            Reaction_time_after_command : Bool := TRUE;   // Start reaction time after command or after shotend
            Spare_0_2 : Bool := FALSE;
            Spare_0_3 : Bool := FALSE;
            Spare_0_4 : Bool := FALSE;
            Spare_0_5 : Bool := FALSE;
            Spare_0_6 : Bool := FALSE;
            Spare_0_7 : Bool := FALSE;
            Spare_1_0 : Bool := FALSE;
            Spare_1_1 : Bool := FALSE;
            Spare_1_2 : Bool := FALSE;
            Spare_1_3 : Bool := FALSE;
            Spare_1_4 : Bool := FALSE;
            Spare_1_5 : Bool := FALSE;
            Spare_1_6 : Bool := FALSE;
            Spare_1_7 : Bool := FALSE;
            Spare_2_0 : Bool := FALSE;
            Spare_2_1 : Bool := FALSE;
            Vacuum_button_valve_1 : Bool := FALSE;
            Vacuum_button_valve_2 : Bool := FALSE;
            Vacuum_button_valve_3 : Bool := TRUE;
            Vacuum_button_valve_4 : Bool := FALSE;
            Vacuum_button_valve_5 : Bool := FALSE;
            Vacuum_button_valve_6 : Bool := FALSE;
            Spare_3 : Byte := 16#00;
         END_STRUCT;
         Times_WinCap : Struct
            SOD_core_WP : Array[0..32] of Time;   // switch on delay core WP
            SOD_core_BP : Array[0..32] of Time;   // switch on delay core BP
            Duration_core : Array[0..32] of Time;   // duration core without endposition
         END_STRUCT;
         Settings_Special : Struct
            Config_write : Bool := FALSE;
            Config_write_done : Bool := FALSE;
            Spare : Int := 1;
            Core_Input : Array[0..32] of "UDT_CoreSettingsSpecial";
            Core_Type : Array[0..32] of Struct
               NC_WP_1 : Bool;   // Schließerkontakt = 0
               NC_WP_2 : Bool;   // Schließerkontakt = 0
               NC_WP_3 : Bool;   // Schließerkontakt = 0
               NC_WP_4 : Bool;   // Schließerkontakt = 0
               NC_WP_5 : Bool;   // Schließerkontakt = 0
               NC_WP_6 : Bool;   // Schließerkontakt = 0
               Forced_forward_WP : Bool;   // Dauernd angesteuert
               Signal_from_upper_tool_WP : Bool;
               NC_BP_1 : Bool;   // Schließerkontakt = 0
               NC_BP_2 : Bool;   // Schließerkontakt = 0
               NC_BP_3 : Bool;   // Schließerkontakt = 0
               NC_BP_4 : Bool;   // Schließerkontakt = 0
               NC_BP_5 : Bool;   // Schließerkontakt = 0
               NC_BP_6 : Bool;   // Schließerkontakt = 0
               Forced_forward_BP : Bool;   // Dauernd angesteuert
               Signal_from_upper_tool_BP : Bool;
            END_STRUCT;
            Config_I_O : Struct
               Lower_tool_card : Array[1..16] of Bool;   // Karte vorhanden
               Upper_tool_card : Array[1..16] of Bool;   // Karte vorhanden
            END_STRUCT;
         END_STRUCT;
      END_STRUCT;
      Set_flow_seals : Struct
         Warning_Tolerance : Struct   // Warning/Tolerance for each seal
            Warning : Array[0..32] of Int;
            Tolerance : Array[0..32] of Int;
         END_STRUCT;
         Set_flow : Array[0..32] of Int;
         Warning_all : Int;   // Warning for all seals
         Tolerance_all : Int;   // Tolerance for all seals
         Set_flow_all : Int;
         Offset_Flow_1 : Real;
         Offset_Flow_2 : Real;
         Offset_Flow_3 : Real;
         SOD_Seal_test : Time := T#2S;   // Waittime to check seal flow
         Spare_140 : Int;
         Spare_142 : Int;
         Spare_144 : Int;
         Spare_146 : Int;
      END_STRUCT;
   END_STRUCT;
   // Set_times_movement.Time_MC_WP[0] := T#10S;
   // Set_times_movement.Time_MC_WP[1] := T#10S;
   // Set_times_movement.Time_MC_WP[2] := T#10S;
   // Set_times_movement.Time_MC_WP[3] := T#10S;
   // Set_times_movement.Time_MC_WP[4] := T#10S;
   // Set_times_movement.Time_MC_WP[5] := T#10S;
   // Set_times_movement.Time_MC_WP[6] := T#10S;
   // Set_times_movement.Time_MC_WP[7] := T#10S;
   // Set_times_movement.Time_MC_WP[8] := T#10S;
   // Set_times_movement.Time_MC_WP[9] := T#10S;
   // Set_times_movement.Time_MC_WP[10] := T#10S;
   // Set_times_movement.Time_MC_WP[11] := T#10S;
   // Set_times_movement.Time_MC_WP[12] := T#10S;
   // Set_times_movement.Time_MC_WP[13] := T#10S;
   // Set_times_movement.Time_MC_WP[14] := T#10S;
   // Set_times_movement.Time_MC_WP[15] := T#10S;
   // Set_times_movement.Time_MC_WP[16] := T#10S;
   // Set_times_movement.Time_MC_WP[17] := T#10S;
   // Set_times_movement.Time_MC_WP[18] := T#10S;
   // Set_times_movement.Time_MC_WP[19] := T#10S;
   // Set_times_movement.Time_MC_WP[20] := T#10S;
   // Set_times_movement.Time_MC_WP[21] := T#10S;
   // Set_times_movement.Time_MC_WP[22] := T#10S;
   // Set_times_movement.Time_MC_WP[23] := T#10S;
   // Set_times_movement.Time_MC_WP[24] := T#10S;
   // Set_times_movement.Time_MC_WP[25] := T#10S;
   // Set_times_movement.Time_MC_WP[26] := T#10S;
   // Set_times_movement.Time_MC_WP[27] := T#10S;
   // Set_times_movement.Time_MC_WP[28] := T#10S;
   // Set_times_movement.Time_MC_WP[29] := T#10S;
   // Set_times_movement.Time_MC_WP[30] := T#10S;
   // Set_times_movement.Time_MC_WP[31] := T#10S;
   // Set_times_movement.Time_MC_WP[32] := T#10S;
   // Set_times_movement.Time_MC_BP[0] := T#10S;
   // Set_times_movement.Time_MC_BP[1] := T#10S;
   // Set_times_movement.Time_MC_BP[2] := T#10S;
   // Set_times_movement.Time_MC_BP[3] := T#10S;
   // Set_times_movement.Time_MC_BP[4] := T#10S;
   // Set_times_movement.Time_MC_BP[5] := T#10S;
   // Set_times_movement.Time_MC_BP[6] := T#10S;
   // Set_times_movement.Time_MC_BP[7] := T#10S;
   // Set_times_movement.Time_MC_BP[8] := T#10S;
   // Set_times_movement.Time_MC_BP[9] := T#10S;
   // Set_times_movement.Time_MC_BP[10] := T#10S;
   // Set_times_movement.Time_MC_BP[11] := T#10S;
   // Set_times_movement.Time_MC_BP[12] := T#10S;
   // Set_times_movement.Time_MC_BP[13] := T#10S;
   // Set_times_movement.Time_MC_BP[14] := T#10S;
   // Set_times_movement.Time_MC_BP[15] := T#10S;
   // Set_times_movement.Time_MC_BP[16] := T#10S;
   // Set_times_movement.Time_MC_BP[17] := T#10S;
   // Set_times_movement.Time_MC_BP[18] := T#10S;
   // Set_times_movement.Time_MC_BP[19] := T#10S;
   // Set_times_movement.Time_MC_BP[20] := T#10S;
   // Set_times_movement.Time_MC_BP[21] := T#10S;
   // Set_times_movement.Time_MC_BP[22] := T#10S;
   // Set_times_movement.Time_MC_BP[23] := T#10S;
   // Set_times_movement.Time_MC_BP[24] := T#10S;
   // Set_times_movement.Time_MC_BP[25] := T#10S;
   // Set_times_movement.Time_MC_BP[26] := T#10S;
   // Set_times_movement.Time_MC_BP[27] := T#10S;
   // Set_times_movement.Time_MC_BP[28] := T#10S;
   // Set_times_movement.Time_MC_BP[29] := T#10S;
   // Set_times_movement.Time_MC_BP[30] := T#10S;
   // Set_times_movement.Time_MC_BP[31] := T#10S;
   // Set_times_movement.Time_MC_BP[32] := T#10S;
   // Set_times_movement.Time_MLD_WP[0] := T#10S;
   // Set_times_movement.Time_MLD_WP[1] := T#10S;
   // Set_times_movement.Time_MLD_WP[2] := T#10S;
   // Set_times_movement.Time_MLD_WP[3] := T#10S;
   // Set_times_movement.Time_MLD_WP[4] := T#10S;
   // Set_times_movement.Time_MLD_WP[5] := T#10S;
   // Set_times_movement.Time_MLD_WP[6] := T#10S;
   // Set_times_movement.Time_MLD_WP[7] := T#10S;
   // Set_times_movement.Time_MLD_WP[8] := T#10S;
   // Set_times_movement.Time_MLD_WP[9] := T#10S;
   // Set_times_movement.Time_MLD_WP[10] := T#10S;
   // Set_times_movement.Time_MLD_WP[11] := T#10S;
   // Set_times_movement.Time_MLD_WP[12] := T#10S;
   // Set_times_movement.Time_MLD_WP[13] := T#10S;
   // Set_times_movement.Time_MLD_WP[14] := T#10S;
   // Set_times_movement.Time_MLD_WP[15] := T#10S;
   // Set_times_movement.Time_MLD_WP[16] := T#10S;
   // Set_times_movement.Time_MLD_WP[17] := T#10S;
   // Set_times_movement.Time_MLD_WP[18] := T#10S;
   // Set_times_movement.Time_MLD_WP[19] := T#10S;
   // Set_times_movement.Time_MLD_WP[20] := T#10S;
   // Set_times_movement.Time_MLD_WP[21] := T#10S;
   // Set_times_movement.Time_MLD_WP[22] := T#10S;
   // Set_times_movement.Time_MLD_WP[23] := T#10S;
   // Set_times_movement.Time_MLD_WP[24] := T#10S;
   // Set_times_movement.Time_MLD_WP[25] := T#10S;
   // Set_times_movement.Time_MLD_WP[26] := T#10S;
   // Set_times_movement.Time_MLD_WP[27] := T#10S;
   // Set_times_movement.Time_MLD_WP[28] := T#10S;
   // Set_times_movement.Time_MLD_WP[29] := T#10S;
   // Set_times_movement.Time_MLD_WP[30] := T#10S;
   // Set_times_movement.Time_MLD_WP[31] := T#10S;
   // Set_times_movement.Time_MLD_WP[32] := T#10S;
   // Set_times_movement.Time_MLD_BP[0] := T#10S;
   // Set_times_movement.Time_MLD_BP[1] := T#10S;
   // Set_times_movement.Time_MLD_BP[2] := T#10S;
   // Set_times_movement.Time_MLD_BP[3] := T#10S;
   // Set_times_movement.Time_MLD_BP[4] := T#10S;
   // Set_times_movement.Time_MLD_BP[5] := T#10S;
   // Set_times_movement.Time_MLD_BP[6] := T#10S;
   // Set_times_movement.Time_MLD_BP[7] := T#10S;
   // Set_times_movement.Time_MLD_BP[8] := T#10S;
   // Set_times_movement.Time_MLD_BP[9] := T#10S;
   // Set_times_movement.Time_MLD_BP[10] := T#10S;
   // Set_times_movement.Time_MLD_BP[11] := T#10S;
   // Set_times_movement.Time_MLD_BP[12] := T#10S;
   // Set_times_movement.Time_MLD_BP[13] := T#10S;
   // Set_times_movement.Time_MLD_BP[14] := T#10S;
   // Set_times_movement.Time_MLD_BP[15] := T#10S;
   // Set_times_movement.Time_MLD_BP[16] := T#10S;
   // Set_times_movement.Time_MLD_BP[17] := T#10S;
   // Set_times_movement.Time_MLD_BP[18] := T#10S;
   // Set_times_movement.Time_MLD_BP[19] := T#10S;
   // Set_times_movement.Time_MLD_BP[20] := T#10S;
   // Set_times_movement.Time_MLD_BP[21] := T#10S;
   // Set_times_movement.Time_MLD_BP[22] := T#10S;
   // Set_times_movement.Time_MLD_BP[23] := T#10S;
   // Set_times_movement.Time_MLD_BP[24] := T#10S;
   // Set_times_movement.Time_MLD_BP[25] := T#10S;
   // Set_times_movement.Time_MLD_BP[26] := T#10S;
   // Set_times_movement.Time_MLD_BP[27] := T#10S;
   // Set_times_movement.Time_MLD_BP[28] := T#10S;
   // Set_times_movement.Time_MLD_BP[29] := T#10S;
   // Set_times_movement.Time_MLD_BP[30] := T#10S;
   // Set_times_movement.Time_MLD_BP[31] := T#10S;
   // Set_times_movement.Time_MLD_BP[32] := T#10S;
   // Set_times_seals.SOD_seal[0] := T#2S;
   // Set_times_seals.SOD_seal[1] := T#2S;
   // Set_times_seals.SOD_seal[2] := T#2S;
   // Set_times_seals.SOD_seal[3] := T#2S;
   // Set_times_seals.SOD_seal[4] := T#2S;
   // Set_times_seals.SOD_seal[5] := T#2S;
   // Set_times_seals.SOD_seal[6] := T#2S;
   // Set_times_seals.SOD_seal[7] := T#2S;
   // Set_times_seals.SOD_seal[8] := T#2S;
   // Set_times_seals.SOD_seal[9] := T#2S;
   // Set_times_seals.SOD_seal[10] := T#2S;
   // Set_times_seals.SOD_seal[11] := T#2S;
   // Set_times_seals.SOD_seal[12] := T#2S;
   // Set_times_seals.SOD_seal[13] := T#2S;
   // Set_times_seals.SOD_seal[14] := T#2S;
   // Set_times_seals.SOD_seal[15] := T#2S;
   // Set_times_seals.SOD_seal[16] := T#2S;
   // Set_times_seals.SOD_seal[17] := T#2S;
   // Set_times_seals.SOD_seal[18] := T#2S;
   // Set_times_seals.SOD_seal[19] := T#2S;
   // Set_times_seals.SOD_seal[20] := T#2S;
   // Set_times_seals.SOD_seal[21] := T#2S;
   // Set_times_seals.SOD_seal[22] := T#2S;
   // Set_times_seals.SOD_seal[23] := T#2S;
   // Set_times_seals.SOD_seal[24] := T#2S;
   // Set_times_seals.SOD_seal[25] := T#2S;
   // Set_times_seals.SOD_seal[26] := T#2S;
   // Set_times_seals.SOD_seal[27] := T#2S;
   // Set_times_seals.SOD_seal[28] := T#2S;
   // Set_times_seals.SOD_seal[29] := T#2S;
   // Set_times_seals.SOD_seal[30] := T#2S;
   // Set_times_seals.SOD_seal[31] := T#2S;
   // Set_times_seals.SOD_seal[32] := T#2S;
   // Set_times_seals.Duration_seal[0] := T#1M_1S;
   // Set_times_seals.Duration_seal[1] := T#1M_1S;
   // Set_times_seals.Duration_seal[2] := T#1M;
   // Set_times_seals.Duration_seal[3] := T#1M;
   // Set_times_seals.Duration_seal[4] := T#1M;
   // Set_times_seals.Duration_seal[5] := T#1M;
   // Set_times_seals.Duration_seal[6] := T#1M;
   // Set_times_seals.Duration_seal[7] := T#1M;
   // Set_times_seals.Duration_seal[8] := T#1M;
   // Set_times_seals.Duration_seal[9] := T#1M;
   // Set_times_seals.Duration_seal[10] := T#1M;
   // Set_times_seals.Duration_seal[11] := T#1M;
   // Set_times_seals.Duration_seal[12] := T#1M;
   // Set_times_seals.Duration_seal[13] := T#1M;
   // Set_times_seals.Duration_seal[14] := T#1M;
   // Set_times_seals.Duration_seal[15] := T#1M;
   // Set_times_seals.Duration_seal[16] := T#1M;
   // Set_times_seals.Duration_seal[17] := T#1M;
   // Set_times_seals.Duration_seal[18] := T#1M;
   // Set_times_seals.Duration_seal[19] := T#1M;
   // Set_times_seals.Duration_seal[20] := T#1M;
   // Set_times_seals.Duration_seal[21] := T#1M;
   // Set_times_seals.Duration_seal[22] := T#1M;
   // Set_times_seals.Duration_seal[23] := T#1M;
   // Set_times_seals.Duration_seal[24] := T#1M;
   // Set_times_seals.Duration_seal[25] := T#1M;
   // Set_times_seals.Duration_seal[26] := T#1M;
   // Set_times_seals.Duration_seal[27] := T#1M;
   // Set_times_seals.Duration_seal[28] := T#1M;
   // Set_times_seals.Duration_seal[29] := T#1M;
   // Set_times_seals.Duration_seal[30] := T#1M;
   // Set_times_seals.Duration_seal[31] := T#1M;
   // Set_times_seals.Duration_seal[32] := T#10S;
   // Set_temperature.Setvalue[0] := 0;
   // Set_temperature.Setvalue[1] := 500;
   // // 1726 more start values not shown
END_TYPE

TYPE "UDT_Mould_functions_1"
VERSION : 0.1
   STRUCT
      MouldMovement01WP : Bool;   // 65: Pusher Windshield WP
      MouldMovement02WP : Bool;   // 66: Pusher Knee Border WP
      MouldMovement03WP : Bool;   // 67: Pusher Frontal Area WP
      MouldMovement04WP : Bool;   // 68: Ejector WP
      MouldMovement05WP : Bool;   // 69: Pusher Stössel WP
      MouldMovement06WP : Bool;   // 70: Flip-Flap WP
      MouldMovement07WP : Bool;   // 71: Safty Locking Knee WP
      MouldMovement08WP : Bool;   // 72: Safty Locking WS WP
      MouldMovement09WP : Bool;   // 73: Vacuum lower mould WP
      MouldMovement10WP : Bool;   // 74: Pusher Airbag WP
      MouldMovement11WP : Bool;   // 75: Pusher DS&PS upper mould WP
      MouldMovement12WP : Bool;   // 76: Vacuum upper mould WP
      MouldMovement13WP : Bool;   // 77: Sensor substrate WP
      MouldMovement14WP : Bool;   // 78: Sensor substrate flamed WP
      MouldMovement15WP : Bool;   // 79: Kernzug 15 AS
      MouldMovement16WP : Bool;   // 80: Kernzug 16 AS
      MouldMovement17WP : Bool;   // 81: Kernzug 17 AS
      MouldMovement18WP : Bool;   // 82: Kernzug 18 AS
      MouldMovement19WP : Bool;   // 83: Kernzug 19 AS
      MouldMovement20WP : Bool;   // 84: Kernzug 20 AS
      MouldMovement21WP : Bool;   // 85: Kernzug 21 AS
      MouldMovement22WP : Bool;   // 86: Kernzug 22 AS
      MouldMovement23WP : Bool;   // 87: Kernzug 23 AS
      MouldMovement24WP : Bool;   // 88: Kernzug 24 AS
      MouldMovement25WP : Bool;   // 89: Kernzug 25 AS
      MouldMovement26WP : Bool;   // 90: Kernzug 26 AS
      MouldMovement27WP : Bool;   // 91: Kernzug 27 AS
      MouldMovement28WP : Bool;   // 92: Kernzug 28 AS
      MouldMovement29WP : Bool;   // 93: Kernzug 29 AS
      MouldMovement30WP : Bool;   // 94: Kernzug 30 AS
      MouldMovement31WP : Bool;   // 95: Kernzug 31 AS
      MouldMovement32WP : Bool;   // 96: Kernzug 32 AS
      MouldMovement01BP : Bool;   // 97: Pusher Windshield BP
      MouldMovement02BP : Bool;   // 98: Pusher Knee Border DS BP
      MouldMovement03BP : Bool;   // 99: Pusher Frontal Area BP
      MouldMovement04BP : Bool;   // 100: Ejector BP
      MouldMovement05BP : Bool;   // 101: Pusher Stössel BP
      MouldMovement06BP : Bool;   // 102: Flip-Flap BP
      MouldMovement07BP : Bool;   // 103: Safty Locking Knee BP
      MouldMovement08BP : Bool;   // 104: Safty Locking WS BP
      MouldMovement09BP : Bool;   // 105: Vacuum lower mould BP
      MouldMovement10BP : Bool;   // 106: Pusher Airbag BP
      MouldMovement11BP : Bool;   // 107: Pusher DS&PS upper mould BP
      MouldMovement12BP : Bool;   // 108: Vacuum upper mould BP
      MouldMovement13BP : Bool;   // 109: Sensor substrate BP
      MouldMovement14BP : Bool;   // 110: Sensor substrate flamed BP
      MouldMovement15BP : Bool;   // 111: Kernzug 15 GS
      MouldMovement16BP : Bool;   // 112: Kernzug 16 GS
      MouldMovement17BP : Bool;   // 113: Kernzug 17 GS
      MouldMovement18BP : Bool;   // 114: Kernzug 18 GS
      MouldMovement19BP : Bool;   // 115: Kernzug 19 GS
      MouldMovement20BP : Bool;   // 116: Kernzug 20 GS
      MouldMovement21BP : Bool;   // 117: Kernzug 21 GS
      MouldMovement22BP : Bool;   // 118: Kernzug 22 GS
      MouldMovement23BP : Bool;   // 119: Kernzug 23 GS
      MouldMovement24BP : Bool;   // 120: Kernzug 24 GS
      MouldMovement25BP : Bool;   // 121: Kernzug 25 GS
      MouldMovement26BP : Bool;   // 122: Kernzug 26 GS
      MouldMovement27BP : Bool;   // 123: Kernzug 27 GS
      MouldMovement28BP : Bool;   // 124: Kernzug 28 GS
      MouldMovement29BP : Bool;   // 125: Kernzug 29 GS
      MouldMovement30BP : Bool;   // 126: Kernzug 30 GS
      MouldMovement31BP : Bool;   // 127: Kernzug 31 GS
      MouldMovement32BP : Bool;   // 128: Kernzug 32 GS
   END_STRUCT;
END_TYPE

TYPE "UDT_Tool_Inputs_type_1"
VERSION : 0.1
   STRUCT
      "Lower Mould" : Struct
         "2A1" : Struct
            I_Pusher_Windshield_DS_WP : Bool := FALSE;   // 0.0
            I_Pusher_Windshield_DS_BP : Bool := FALSE;   // 0.1
            Reserve_5 : Bool := FALSE;   // 0.2
            Reserve_4 : Bool := FALSE;   // 0.3
            I_Pusher_Knee_Border_DS_WP : Bool := FALSE;   // 0.4
            I_Pusher_Knee_Border_DS_BP : Bool := FALSE;   // 0.5
            Reserve_3 : Bool := FALSE;   // 0.6
            Reserve_2 : Bool := FALSE;   // 0.7
            I_Pusher_Frontal_Area_DS_WP : Bool := FALSE;   // 1.0
            I_Pusher_Frontal_Area_DS_BP : Bool := FALSE;   // 1.1
            I_Pusher_Frontal_Area_PS_WP : Bool := FALSE;   // 1.2
            I_Pusher_Frontal_Area_PS_BP : Bool := FALSE;   // 1.3
            I_Ejector_WP : Bool := FALSE;   // 1.4
            I_Ejector_BP : Bool := FALSE;   // 1.5
            "I_Flip-Flap_WP" : Bool := FALSE;   // 1.6
            Reserve_1 : Bool := FALSE;   // 1.7
         END_STRUCT;
         "2A2" : Struct
            I_Safty_Locking_Knee_DS_WP : Bool := FALSE;   // 0.0
            I_Safty_Locking_Knee_DS_BP : Bool := FALSE;   // 0.1
            I_Safty_Locking_Knee_PS_WP : Bool := FALSE;   // 0.2
            I_Safty_Locking_Knee_PS_BP : Bool := FALSE;   // 0.3
            I_Safty_Locking_WS_DS_WP : Bool := FALSE;   // 0.4
            I_Safty_Locking_WS_DS_BP : Bool := FALSE;   // 0.5
            I_Safty_Locking_WS_PS_WP : Bool := FALSE;   // 0.6
            I_Safty_Locking_WS_PS_BP : Bool := FALSE;   // 0.7
            "I_Vacuum monitor" : Bool := FALSE;   // 1.0
            Element_2 : Bool := FALSE;   // 1.1
            Element_1 : Bool := FALSE;   // 1.2
            Element_4 : Bool := FALSE;   // 1.3
            Reserve_2 : Bool := FALSE;   // 1.4
            Reserve_3 : Bool := FALSE;   // 1.5
            Reserve_4 : Bool := FALSE;   // 1.6
            Reserve_5 : Bool := FALSE;   // 1.7
         END_STRUCT;
         "2A3" : Struct
            I_Palm_Switch_Vacuum_on : Bool := FALSE;   // 0.0
            I_Illuminated_Key_Vacuum1_off : Bool := FALSE;   // 0.1
            I_Illuminated_Key_Vacuum2_off : Bool := FALSE;   // 0.2
            I_Illuminated_Key_Vacuum3_off : Bool := FALSE;   // 0.3
            Element_3 : Bool := FALSE;   // 0.4
            Element_1 : Bool := FALSE;   // 0.5
            I_PB_Seal_Test_2bar : Bool := FALSE;   // 0.6
            I_2_Hand_active : Bool := FALSE;   // 0.7
            "I_Code_Bit1_(1)" : Bool := FALSE;   // 1.0
            "I_Code_Bit2_(2)" : Bool := FALSE;   // 1.1
            "I_Code_Bit3_(4)" : Bool := FALSE;   // 1.2
            "I_Code_Bit4_(8)" : Bool := FALSE;   // 1.3
            "I_Code_Bit5_(16)" : Bool := FALSE;   // 1.4
            "I_Code_Bit6_(32)" : Bool := FALSE;   // 1.5
            "I_Code_Bit7_(64)" : Bool := FALSE;   // 1.6
            "I_Code_Bit8_(128)" : Bool := FALSE;   // 1.7
         END_STRUCT;
      END_STRUCT;
      "Upper Mould" : Struct
         "46A1" : Struct
            I_Pusher_Airbag_WP : Bool := FALSE;   // 0.0
            I_Pusher_Airbag_BP : Bool := FALSE;   // 0.1
            I_Pusher_DS_WP : Bool := FALSE;   // 0.2
            I_Pusher_DS_BP : Bool := FALSE;   // 0.3
            I_Pusher_PS_WP : Bool := FALSE;   // 0.4
            I_Pusher_PS_BP : Bool := FALSE;   // 0.5
            Element_1 : Bool := FALSE;   // 0.6
            Element_2 : Bool := FALSE;   // 0.7
            I_Vacuum_Motitor : Bool := FALSE;   // 1.0
            I_Sensor_insert : Bool := FALSE;   // 1.1
            I_Sensor_flamed : Bool := FALSE;   // 1.2
            "I_Illuminated Key_Vacuum_off" : Bool := FALSE;   // 1.3
            Element_3 : Bool := FALSE;   // 1.4
            Element_4 : Bool := FALSE;   // 1.5
            Reserve_54 : Bool := FALSE;   // 1.6
            Reserve_55 : Bool := FALSE;   // 1.7
         END_STRUCT;
      END_STRUCT;
   END_STRUCT;
END_TYPE

TYPE "UDT1500_ShotResultToMC"
VERSION : 0.1
   STRUCT
      Data_from_MC : Struct
         Struct01 : Struct
            Data_read : Bool;   // Mouldcarrier has read the shot data
            SPARE_00 : Bool;
            SPARE_01 : Bool;
            SPARE_02 : Bool;
            SPARE_03 : Bool;
            SPARE_04 : Bool;
            SPARE_05 : Bool;
            SPARE_06 : Bool;
            SPARE_07 : Bool;
            SPARE_08 : Bool;
            SPARE_09 : Bool;
            SPARE_10 : Bool;
            SPARE_11 : Bool;
            SPARE_12 : Bool;
            SPARE_13 : Bool;
            SPARE_14 : Bool;
         END_STRUCT;
      END_STRUCT;
      Date_to_MC : Struct
         Struct01 : Struct   // 128 Byte Bereich
            New_Data : Bool;   // Shot Data is now available
            SPARE_00 : Bool;
            SPARE_01 : Bool;
            SPARE_02 : Bool;
            SPARE_03 : Bool;
            SPARE_04 : Bool;
            SPARE_05 : Bool;
            SPARE_06 : Bool;
            FLT_Shottime : Bool;   // Shottime is outside of the tolerance
            FLT_Flowrate_C1 : Bool;   // Flowrate of C1 is outside of the tolerance
            FLT_Flowrate_C2 : Bool;   // Flowrate of C2 is outside of the tolerance
            FLT_PressureMH_C1 : Bool;   // Pressure of C1 at the MH is outside of the tolerance
            FLT_PressureMH_C2 : Bool;   // Pressure of C2 at the MH is outside of the tolerance
            FLT_TempMH_C1 : Bool;   // Temperature of C1 at the MH is outside of the tolerance
            FLT_TempMH_C2 : Bool;   // Temperature of C2 at the MH is outside of the tolerance
            FLT_TempTank_C1 : Bool;   // Temperature of C1 at the tank is outside of the tolerance
            FLT_TempTank_C2 : Bool;   // Temperature of C2 at the tank is outside of the tolerance
            SPARE_07 : Bool;
            SPARE_08 : Bool;
            SPARE_09 : Bool;
            SPARE_10 : Bool;
            SPARE_11 : Bool;
            SPARE_12 : Bool;
            SPARE_13 : Bool;
            SPARE_14 : Bool;
            SPARE_15 : Bool;
            SPARE_16 : Bool;
            SPARE_17 : Bool;
            SPARE_18 : Bool;
            SPARE_19 : Bool;
            SPARE_20 : Bool;
            SPARE_21 : Bool;
            MH_No : Int;   // Number of the MH at the last shot (1 - 16)
            Foam_No : Int;   // Number of foaming program at the last shot (1 - 1000)
            MC_No : Int;
            SPARE_22 : Int;
            Rob_MoveTime : DInt;   // Moving - time of the roboter (1/1 [ms])
            ShotTime_Tol_plus : DInt;   // Tolerance of the shottime (plus) at the last shot (1/1 [ms])
            ShotTime_Setvalue : DInt;   // Setvalue of the shottime at the last shot (1/1 [ms])
            ShotTime_Actvalue : DInt;   // Actual value of the shottime at the last shot (1/1 [ms])
            ShotTime_Tol_minus : DInt;   // Tolerance of the shottime (minus) at the last shot (1/1 [ms])
            ShotWeight_Setvalue : DInt;
            ShotWeight_Actvalue : DInt;
            Flowrate_C1_Tol_plus : DInt;   // Tolerance of the flowrate (plus) at the last shot (1/10 [g/s])
            Flowrate_C1_Setvalue : DInt;   // Setvalue of the flowrate at the last shot (1/10 [g/s])
            Flowrate_C1_Actvalue : DInt;   // Actual value of the flowrate at the last shot (1/10 [g/s])
            Flowrate_C1_Tol_minus : DInt;   // Tolerance of the flowrate (minus) at the last shot (1/10 [g/s])
            Flowrate_C2_Tol_plus : DInt;   // Tolerance of the flowrate (plus) at the last shot (1/10 [g/s])
            Flowrate_C2_Setvalue : DInt;   // Setvalue of the flowrate at the last shot (1/10 [g/s])
            Flowrate_C2_Actvalue : DInt;   // Actual value of the flowrate at the last shot (1/10 [g/s])
            Flowrate_C2_Tol_minus : DInt;   // Tolerance of the flowrate (minus) at the last shot (1/10 [g/s])
            PressureMH_C1_Tol_plus : DInt;   // Tolerance of the pressure of C1 at the MH (plus) at the last shot (1/10 [bar])
            PressureMH_C1_Setvalue : DInt;   // Setvalue of the pressure of C1 at the MH at the last shot (1/10 [bar])
            PressureMH_C1_Actvalue : DInt;   // Actual value of the pressure of C1 at the MH at the last shot (1/10 [bar])
            PressureMH_C1_Tol_minus : DInt;   // Tolerance of the pressure of C1 at the MH(minus) at the last shot (1/10 [bar])
            PressureMH_C2_Tol_plus : DInt;   // Tolerance of the pressure of C2 at the MH (plus) at the last shot (1/10 [bar])
            PressureMH_C2_Setvalue : DInt;   // Setvalue of the pressure of C2 at the MH at the last shot (1/10 [bar])
            PressureMH_C2_Actvalue : DInt;   // Actual value of the pressure of C2 at the MH at the last shot (1/10 [bar])
            PressureMH_C2_Tol_minus : DInt;   // Tolerance of the pressure of C2 at the MH(minus) at the last shot (1/10 [bar])
            TempMH_C1_Tol_plus : DInt;   // Tolerance of the temp. of C1 at the MH (plus) at the last shot (1/10 [°C])
            TempMH_C1_Setvalue : DInt;   // Setvalue of the temp. of C1 at the MH at the last shot (1/10 [°C])
            TempMH_C1_Actvalue : DInt;   // Actual value of the temp. of C1 at the MH at the last shot (1/10 [°C])
            TempMH_C1_Tol_minus : DInt;   // Tolerance of the temp. of C1 at the MH(minus) at the last shot (1/10 [°C])
            TempMH_C2_Tol_plus : DInt;   // Tolerance of the temp. of C2 at the MH (plus) at the last shot (1/10 [°C])
            TempMH_C2_Setvalue : DInt;   // Setvalue of the temp. of C2 at the MH at the last shot (1/10 [°C])
         END_STRUCT;
         Struct02 : Struct   // 64 Byte Bereich
            TempMH_C2_Actvalue : DInt;   // Actual value of the temp. of C2 at the MH at the last shot (1/10 [°C])
            TempMH_C2_Tol_minus : DInt;   // Tolerance of the temp. of C2 at the MH(minus) at the last shot (1/10 [°C])
            TempTank_C1_Tol_plus : DInt;   // Tolerance of the temp. of C1 at the tank(plus) at the last shot (1/10 [°C])
            TempTank_C1_Setvalue : DInt;   // Setvalue of the temp. of C1 at the tank at the last shot (1/10 [°C])
            TempTank_C1_Actvalue : DInt;   // Actual value of the temp. of C1 at the tank at the last shot (1/10 [°C])
            TempTank_C1_Tol_minus : DInt;   // Tolerance of the temp. of C1 at the tank(minus) at the last shot (1/10 [°C])
            TempTank_C2_Tol_plus : DInt;   // Tolerance of the temp. of C2 at the tank (plus) at the last shot (1/10 [°C])
            TempTank_C2_Setvalue : DInt;   // Setvalue of the temp. of C2 at the tank at the last shot (1/10 [°C])
            TempTank_C2_Actvalue : DInt;   // Actual value of the temp. of C2 at the tank at the last shot (1/10 [°C])
            TempTank_C2_Tol_minus : DInt;   // Tolerance of the temp. of C2 at the tank (minus) at the last shot (1/10 [°C])
            SPARE_23 : DInt;
            SPARE_24 : DInt;
            SPARE_25 : DInt;
            SPARE_26 : DInt;
            SPARE_27 : DInt;
            SPARE_28 : DInt;
         END_STRUCT;
      END_STRUCT;
   END_STRUCT;
END_TYPE

TYPE "UDT_Seg_input"
VERSION : 0.1
   STRUCT
      I_spare_2x0_0 : Bool;
      I_PS_down : Bool;   // Parallelstroke in lower position
      I_P_okay : Bool;   // Airpressure okay
      I_aircushion_front_down : Bool;   // Aircushion front down
      I_spare_2x0_4 : Bool;
      I_P_aircushion_down : Bool;   // Pressure switch aircushion down
      I_P_aircushion_up : Bool;   // Pressure switch aircushion up
      I_spare_2x0_7 : Bool;
      I_L_bold_unlocked : Bool;   // Left bold lower/upper plate unlocked
      I_L_bold_locked : Bool;   // Left bold lower/upper plate locked
      I_R_bold_unlocked : Bool;   // Right bold lower/upper plate unlocked
      I_R_bold_locked : Bool;   // Right bold lower/upper plate locked
      I_Reference_position_PS : Bool;   // Sensor reference position parallel stroke
      I_spare_2x1_5 : Bool;
      I_spare_2x1_6 : Bool;
      I_spare_2x1_7 : Bool;
      I_L_U_Safetybold_unlocked : Bool;   // Left upper safety bold unlocked
      I_L_U_Safetybold_locked : Bool;   // Left upper safety bold locked
      I_L_L_Safetybold_unlocked : Bool;   // Left lower safety bold unlocked
      I_L_L_Safetybold_locked : Bool;   // Left lower safety bold locked
      I_R_U_Safetybold_unlocked : Bool;   // Right upper safety bold unlocked
      I_R_U_Safetybold_locked : Bool;   // Right upper safety bold locked
      I_R_L_Safetybold_unlocked : Bool;   // Right lower safety bold unlocked
      I_R_L_Safetybold_locked : Bool;   // Right lower safety bold locked
      I_UMP_Safetybold_1_unlocked : Bool;   // safety bold 1 upper mold plate unlocked
      I_UMP_Safetybold_1_locked : Bool;   // safety bold 1 upper mold plate locked
      I_UMP_Safetybold_2_unlocked : Bool;   // safety bold 2 upper mold plate unlocked
      I_UMP_Safetybold_2_locked : Bool;   // safety bold 2 upper mold plate locked
      I_Reference_position_UMP : Bool;   // Sensor reference position upper mold plate
      I_Reference_position_LMP : Bool;   // Sensor reference position lower mold plate
      I_spare_2x3_6 : Bool;
      I_spare_2x3_7 : Bool;
      I_spare_2x4_0 : Bool;
      I_spare_2x4_1 : Bool;
      I_spare_2x4_2 : Bool;
      I_spare_2x4_3 : Bool;
      I_Reference_position_frame : Bool;   // Sensor reference position frame
      I_spare_2x4_5 : Bool;
      I_spare_2x4_6 : Bool;
      I_spare_2x4_7 : Bool;
      I_MldLckLP_l_locked : Bool;   // Left bold tool change lower plate locked
      I_MldLckLP_r_locked : Bool;   // Right bold tool change lower plate locked
      I_spare_2x5_2 : Bool;
      I_spare_2x5_3 : Bool;
      I_MldLckUP_l_unlocked : Bool;   // Left bold tool change upper plate unlocked
      I_MldLckUP_l_locked : Bool;   // Left bold tool change upper plate locked
      I_MldLckUP_r_unlocked : Bool;   // Right bold tool change upper plate unlocked
      I_MldLckUP_r_locked : Bool;   // Right bold tool change upper plate locked
      I_Tool_LP_Code0 : Bool;   // Input Toolcode lower plate Bit 0
      I_Tool_LP_Code1 : Bool;   // Input Toolcode lower plate Bit 1
      I_Tool_LP_Code2 : Bool;   // Input Toolcode lower plate Bit 2
      I_Tool_LP_Code3 : Bool;   // Input Toolcode lower plate Bit 3
      I_Tool_UP_Code0 : Bool;   // Input Toolcode upper plate Bit 0
      I_Tool_UP_Code1 : Bool;   // Input Toolcode upper plate Bit 1
      I_Tool_UP_Code2 : Bool;   // Input Toolcode upper plate Bit 2
      I_Tool_UP_Code3 : Bool;   // Input Toolcode upper plate Bit 3
   END_STRUCT;
END_TYPE

TYPE "UDT_CoreHydraulic"
VERSION : 0.0
   STRUCT
      FLT_motor_protection_hydraulic : Bool;   // Störung: Der Versorgungsspanung oder des Motorschutzes des Hydraulikaggregates
      FLT_motor_protection_ventilation : Bool;   // Störung: Der Versorgungsspanung oder des Motorschutzes des Ventilators
      FLT_min_level_oil : Bool;   // Störung: Der minimale Füllstand des Hydrauliköls wurde unterschritten
      WRN_max_temp : Bool;   // Warnung: Die eingestellte max. Temperatur wurde überschritten
      FLT_max_temp : Bool;   // Störung: Die eingestellte max. Temperatur wurde länger als 5 Min. überschritten
      FLT_pressure_reached : Bool;   // Störung: Der nötige Druck wird innerhalb der festgelegten Zeit nicht erreicht
      Spare_1_5 : Bool;
      Spare_1_6 : Bool;
      Request_motor : Bool;   // Hydraulikmotor einschalten
      Request_motor_done : Bool;   // Der Anlauf des Hydraulikmotors ist beendet
      Hydraulic_okay : Bool;   // Die Hydraulik läuft und der eingestellte Betriebsdruck wurde erreicht
      Flag_T_ON : Bool;   // Flankenhilfsmerker zum Ein- Ausschalten des Hydraulikmotors
      General_FLT : Bool;   // Es steht eine Störung an, der Motor wird abgeschaltet
      OUT_motor_net : Bool;   // Ansteuerung des Netz- Schützes des Hydraulik- Motors
      OUT_Pressure_valve : Bool;   // Ansteuerung des Druckaufbauventils der Mischkopfhydraulik
      OUT_Ventilation : Bool;   // Ansteuerung des Ventilators für die Ölkühlung
   END_STRUCT;
END_TYPE

TYPE "UDT_State_MC"
VERSION : 0.1
   STRUCT
      Movement : Struct
         RequestFromOP : "UDT_Actions";
         Request : "UDT_Actions";
         Command : "UDT_Actions";
         Valve : "UDT_Actions";
         End : "UDT_Actions";
      END_STRUCT;
      State : Struct
         Tool_No : Byte := B#16#0;
         MC_blocked : Bool := FALSE;
         MC_selected : Bool := FALSE;
         Tool_exists : Bool := FALSE;
         Fault_MC : Bool := FALSE;
         Turnlock : Bool := FALSE;
         Spare_1 : Bool := FALSE;
         Delete_cycle : Bool := FALSE;
         Spare_2 : Bool := FALSE;
         MC_request_foamingcycle : Bool := FALSE;
         Spare_3 : Bool := FALSE;
         Request_degasing : Bool := FALSE;
         Request_homecycle : Bool := FALSE;
         Request_breakcycle : Bool := FALSE;
         Request_toolchangecycle : Bool := FALSE;
         Spare_4 : Bool := FALSE;
         Homeposition_active : Bool := FALSE;
         Homeposition_end : Bool := FALSE;
         Foamingcycle_active : Bool := FALSE;
         Foamingcycle_end : Bool := FALSE;
         MC_was_in_degasing_position : Bool := FALSE;
         Breakposition_active : Bool := FALSE;
         Breakposition_end : Bool := FALSE;
         MC_in_break_position : Bool := FALSE;
         Toolchange_active : Bool := FALSE;
         Toolchange_end : Bool := FALSE;
         Spare_5 : Bool := FALSE;
         Spare_6 : Bool := FALSE;
         MC_Shotpreperation : Bool := FALSE;
         MC_Shotrelease : Bool := FALSE;
         MC_Shotend : Bool := FALSE;
         MC_Shotfault : Bool := FALSE;
         Start_seal_times : Bool := FALSE;
         MC_program_end : Bool := FALSE;
         B_no_foaming : Bool := FALSE;
         MC_cycle_started : Bool := FALSE;
         MC_foamed : Bool := FALSE;
         Reactiontime : Bool := FALSE;
         MC_cycle_running : Bool := FALSE;
         Flag_start_foaming : Bool := FALSE;
         Flag_stop_foaming : Bool := FALSE;
         Spare_7 : Bool := FALSE;
         Spare_8 : Bool := FALSE;
         Spare_9 : Bool := FALSE;
         Spare_10 : Bool := FALSE;
         Spare_11 : Bool := FALSE;
         Spare_12 : Bool := FALSE;
         Spare_13 : Bool := FALSE;
         Spare_14 : Bool := FALSE;
         Spare_15 : Bool := FALSE;
         Flag_TT_not_in_position : Bool := FALSE;
         Spare_16 : Bool := FALSE;
         Release_production : Bool := FALSE;
         Flag_Counter_iO : Bool := FALSE;
         Flag_Counter_niO : Bool := FALSE;
         Spare_17 : Bool := FALSE;
         Spare_18 : Bool := FALSE;
         Spare_19 : Word := W#16#0;
         FM_Haltung_UT : Bool := FALSE;
         Zutrittsfreigabe_von_FT : Bool := FALSE;
         Beflammen_verwerfen : Bool := FALSE;
         Teil_i_O : Bool := FALSE;
         Bedienung_OP177 : Bool := FALSE;
         Zyklus_abbrechen : Bool := FALSE;
         FHM_Vakuum_OT_1 : Bool := FALSE;
         FHM_Vakuum_OT_2 : Bool := FALSE;
         FHM_Vakuum_UT_1 : Bool := FALSE;
         Flanke_Counter_13 : Bool := FALSE;
         Flanke_Counter_12 : Bool := FALSE;
         Flanke_Counter_11 : Bool := FALSE;
         Dichtung_12_Ein : Bool := FALSE;
         Dichtung_11_Ein : Bool := FALSE;
         Dichtung_10_Ein : Bool := FALSE;
         Dichtung_09_Ein : Bool := FALSE;
         Dichtung_01_Ein : Bool := FALSE;
         Dichtung_02_Ein : Bool := FALSE;
         Dichtung_03_Ein : Bool := FALSE;
         Dichtung_04_Ein : Bool := FALSE;
         Dichtung_05_Ein : Bool := FALSE;
         Dichtung_06_Ein : Bool := FALSE;
         Dichtung_07_Ein : Bool := FALSE;
         Dichtung_08_Ein : Bool := FALSE;
         Dichtungen_Aus : Bool := FALSE;
         STG_Warn_Min_Temp_OT : Bool := FALSE;
         STG_Tol_Min_Temp_OT : Bool := FALSE;
         STG_Warn_Max_Temp_OT : Bool := FALSE;
         STG_Tol_Max_Temp_OT : Bool := FALSE;
         HM_Entl_Deckel : Bool := FALSE;
         Flanke_Counter_01 : Bool := FALSE;
         Flanke_Counter_02 : Bool := FALSE;
         Flanke_Counter_03 : Bool := FALSE;
         Flanke_Counter_04 : Bool := FALSE;
         Flanke_Counter_05 : Bool := FALSE;
         Flanke_Counter_06 : Bool := FALSE;
         Flanke_Counter_07 : Bool := FALSE;
         Flanke_Counter_08 : Bool := FALSE;
         Flanke_Counter_09 : Bool := FALSE;
         Flanke_Counter_10 : Bool := FALSE;
         Reserve_18 : Word := W#16#0;
         Reserve_20 : Word := W#16#0;
      END_STRUCT;
   END_STRUCT;
   // Movement.RequestFromOP.MCMovement01WP := FALSE;
   // Movement.RequestFromOP.MCMovement02WP := FALSE;
   // Movement.RequestFromOP.MCMovement03WP := FALSE;
   // Movement.RequestFromOP.MCMovement04WP := FALSE;
   // Movement.RequestFromOP.MCMovement05WP := FALSE;
   // Movement.RequestFromOP.MCMovement06WP := FALSE;
   // Movement.RequestFromOP.MCMovement07WP := FALSE;
   // Movement.RequestFromOP.MCMovement08WP := FALSE;
   // Movement.RequestFromOP.MCMovement09WP := FALSE;
   // Movement.RequestFromOP.MCMovement10WP := FALSE;
   // Movement.RequestFromOP.MCMovement11WP := FALSE;
   // Movement.RequestFromOP.MCMovement12WP := FALSE;
   // Movement.RequestFromOP.MCMovement13WP := FALSE;
   // Movement.RequestFromOP.MCMovement14WP := FALSE;
   // Movement.RequestFromOP.MCMovement15WP := FALSE;
   // Movement.RequestFromOP.MCMovement16WP := FALSE;
   // Movement.RequestFromOP.MCMovement17WP := FALSE;
   // Movement.RequestFromOP.MCMovement18WP := FALSE;
   // Movement.RequestFromOP.MCMovement19WP := FALSE;
   // Movement.RequestFromOP.MCMovement20WP := FALSE;
   // Movement.RequestFromOP.MCMovement21WP := FALSE;
   // Movement.RequestFromOP.MCMovement22WP := FALSE;
   // Movement.RequestFromOP.MCMovement23WP := FALSE;
   // Movement.RequestFromOP.MCMovement24WP := FALSE;
   // Movement.RequestFromOP.MCMovement25WP := FALSE;
   // Movement.RequestFromOP.MCMovement26WP := FALSE;
   // Movement.RequestFromOP.MCMovement27WP := FALSE;
   // Movement.RequestFromOP.MCMovement28WP := FALSE;
   // Movement.RequestFromOP.MCMovement29WP := FALSE;
   // Movement.RequestFromOP.MCMovement30WP := FALSE;
   // Movement.RequestFromOP.MCMovement31WP := FALSE;
   // Movement.RequestFromOP.MCMovement32WP := FALSE;
   // Movement.RequestFromOP.MCMovement01BP := FALSE;
   // Movement.RequestFromOP.MCMovement02BP := FALSE;
   // Movement.RequestFromOP.MCMovement03BP := FALSE;
   // Movement.RequestFromOP.MCMovement04BP := FALSE;
   // Movement.RequestFromOP.MCMovement05BP := FALSE;
   // Movement.RequestFromOP.MCMovement06BP := FALSE;
   // Movement.RequestFromOP.MCMovement07BP := FALSE;
   // Movement.RequestFromOP.MCMovement08BP := FALSE;
   // Movement.RequestFromOP.MCMovement09BP := FALSE;
   // Movement.RequestFromOP.MCMovement10BP := FALSE;
   // Movement.RequestFromOP.MCMovement11BP := FALSE;
   // Movement.RequestFromOP.MCMovement12BP := FALSE;
   // Movement.RequestFromOP.MCMovement13BP := FALSE;
   // Movement.RequestFromOP.MCMovement14BP := FALSE;
   // Movement.RequestFromOP.MCMovement15BP := FALSE;
   // Movement.RequestFromOP.MCMovement16BP := FALSE;
   // Movement.RequestFromOP.MCMovement17BP := FALSE;
   // Movement.RequestFromOP.MCMovement18BP := FALSE;
   // Movement.RequestFromOP.MCMovement19BP := FALSE;
   // Movement.RequestFromOP.MCMovement20BP := FALSE;
   // Movement.RequestFromOP.MCMovement21BP := FALSE;
   // Movement.RequestFromOP.MCMovement22BP := FALSE;
   // Movement.RequestFromOP.MCMovement23BP := FALSE;
   // Movement.RequestFromOP.MCMovement24BP := FALSE;
   // Movement.RequestFromOP.MCMovement25BP := FALSE;
   // Movement.RequestFromOP.MCMovement26BP := FALSE;
   // Movement.RequestFromOP.MCMovement27BP := FALSE;
   // Movement.RequestFromOP.MCMovement28BP := FALSE;
   // Movement.RequestFromOP.MCMovement29BP := FALSE;
   // Movement.RequestFromOP.MCMovement30BP := FALSE;
   // Movement.RequestFromOP.MCMovement31BP := FALSE;
   // Movement.RequestFromOP.MCMovement32BP := FALSE;
   // Movement.RequestFromOP.MouldMovement01WP := FALSE;
   // Movement.RequestFromOP.MouldMovement02WP := FALSE;
   // Movement.RequestFromOP.MouldMovement03WP := FALSE;
   // Movement.RequestFromOP.MouldMovement04WP := FALSE;
   // Movement.RequestFromOP.MouldMovement05WP := FALSE;
   // Movement.RequestFromOP.MouldMovement06WP := FALSE;
   // Movement.RequestFromOP.MouldMovement07WP := FALSE;
   // Movement.RequestFromOP.MouldMovement08WP := FALSE;
   // Movement.RequestFromOP.MouldMovement09WP := FALSE;
   // Movement.RequestFromOP.MouldMovement10WP := FALSE;
   // Movement.RequestFromOP.MouldMovement11WP := FALSE;
   // Movement.RequestFromOP.MouldMovement12WP := FALSE;
   // Movement.RequestFromOP.MouldMovement13WP := FALSE;
   // Movement.RequestFromOP.MouldMovement14WP := FALSE;
   // Movement.RequestFromOP.MouldMovement15WP := FALSE;
   // Movement.RequestFromOP.MouldMovement16WP := FALSE;
   // Movement.RequestFromOP.MouldMovement17WP := FALSE;
   // Movement.RequestFromOP.MouldMovement18WP := FALSE;
   // Movement.RequestFromOP.MouldMovement19WP := FALSE;
   // Movement.RequestFromOP.MouldMovement20WP := FALSE;
   // Movement.RequestFromOP.MouldMovement21WP := FALSE;
   // Movement.RequestFromOP.MouldMovement22WP := FALSE;
   // Movement.RequestFromOP.MouldMovement23WP := FALSE;
   // Movement.RequestFromOP.MouldMovement24WP := FALSE;
   // Movement.RequestFromOP.MouldMovement25WP := FALSE;
   // Movement.RequestFromOP.MouldMovement26WP := FALSE;
   // Movement.RequestFromOP.MouldMovement27WP := FALSE;
   // Movement.RequestFromOP.MouldMovement28WP := FALSE;
   // Movement.RequestFromOP.MouldMovement29WP := FALSE;
   // Movement.RequestFromOP.MouldMovement30WP := FALSE;
   // Movement.RequestFromOP.MouldMovement31WP := FALSE;
   // Movement.RequestFromOP.MouldMovement32WP := FALSE;
   // Movement.RequestFromOP.MouldMovement01BP := FALSE;
   // Movement.RequestFromOP.MouldMovement02BP := FALSE;
   // Movement.RequestFromOP.MouldMovement03BP := FALSE;
   // Movement.RequestFromOP.MouldMovement04BP := FALSE;
   // Movement.RequestFromOP.MouldMovement05BP := FALSE;
   // Movement.RequestFromOP.MouldMovement06BP := FALSE;
   // Movement.RequestFromOP.MouldMovement07BP := FALSE;
   // Movement.RequestFromOP.MouldMovement08BP := FALSE;
   // Movement.RequestFromOP.MouldMovement09BP := FALSE;
   // Movement.RequestFromOP.MouldMovement10BP := FALSE;
   // Movement.RequestFromOP.MouldMovement11BP := FALSE;
   // Movement.RequestFromOP.MouldMovement12BP := FALSE;
   // Movement.RequestFromOP.MouldMovement13BP := FALSE;
   // Movement.RequestFromOP.MouldMovement14BP := FALSE;
   // Movement.RequestFromOP.MouldMovement15BP := FALSE;
   // Movement.RequestFromOP.MouldMovement16BP := FALSE;
   // Movement.RequestFromOP.MouldMovement17BP := FALSE;
   // Movement.RequestFromOP.MouldMovement18BP := FALSE;
   // Movement.RequestFromOP.MouldMovement19BP := FALSE;
   // Movement.RequestFromOP.MouldMovement20BP := FALSE;
   // Movement.RequestFromOP.MouldMovement21BP := FALSE;
   // Movement.RequestFromOP.MouldMovement22BP := FALSE;
   // Movement.RequestFromOP.MouldMovement23BP := FALSE;
   // Movement.RequestFromOP.MouldMovement24BP := FALSE;
   // Movement.RequestFromOP.MouldMovement25BP := FALSE;
   // Movement.RequestFromOP.MouldMovement26BP := FALSE;
   // Movement.RequestFromOP.MouldMovement27BP := FALSE;
   // Movement.RequestFromOP.MouldMovement28BP := FALSE;
   // Movement.RequestFromOP.MouldMovement29BP := FALSE;
   // Movement.RequestFromOP.MouldMovement30BP := FALSE;
   // Movement.RequestFromOP.MouldMovement31BP := FALSE;
   // Movement.RequestFromOP.MouldMovement32BP := FALSE;
   // Movement.RequestFromOP.ShotPreparation := FALSE;
   // Movement.RequestFromOP.ShotEnable := FALSE;
   // Movement.RequestFromOP.ShotEnd := FALSE;
   // Movement.RequestFromOP.StartReactionTime := FALSE;
   // Movement.RequestFromOP.WaitReactionTime := FALSE;
   // Movement.RequestFromOP.Spare134 := FALSE;
   // Movement.RequestFromOP.Spare135 := FALSE;
   // Movement.RequestFromOP.Spare136 := FALSE;
   // Movement.RequestFromOP.Spare137 := FALSE;
   // Movement.RequestFromOP.Spare138 := FALSE;
   // Movement.RequestFromOP.WaitTime1 := FALSE;
   // Movement.RequestFromOP.WaitTime2 := FALSE;
   // Movement.RequestFromOP.WaitTime3 := FALSE;
   // Movement.RequestFromOP.WaitTime4 := FALSE;
   // Movement.RequestFromOP.WaitTime5 := FALSE;
   // Movement.RequestFromOP.WaitTime6 := FALSE;
   // Movement.RequestFromOP.StopCycle := FALSE;
   // Movement.RequestFromOP.Spare146 := FALSE;
   // Movement.RequestFromOP.NoFaultGroup1 := FALSE;
   // Movement.RequestFromOP.SafetyOk := FALSE;
   // Movement.RequestFromOP.StartWatch := FALSE;
   // Movement.RequestFromOP.StopWatch := FALSE;
   // Movement.RequestFromOP.Spare151 := FALSE;
   // Movement.RequestFromOP.Spare152 := FALSE;
   // Movement.RequestFromOP.Spare153 := FALSE;
   // Movement.RequestFromOP.Spare154 := FALSE;
   // Movement.RequestFromOP.Spare155 := FALSE;
   // Movement.RequestFromOP.Spare156 := FALSE;
   // Movement.RequestFromOP.Set_access_release := FALSE;
   // Movement.RequestFromOP.Reset_access_release := FALSE;
   // Movement.RequestFromOP.RobotOutOfMC := FALSE;
   // Movement.RequestFromOP.EndOfProgram := FALSE;
   // Movement.Request.MCMovement01WP := FALSE;
   // Movement.Request.MCMovement02WP := FALSE;
   // Movement.Request.MCMovement03WP := FALSE;
   // Movement.Request.MCMovement04WP := FALSE;
   // Movement.Request.MCMovement05WP := FALSE;
   // Movement.Request.MCMovement06WP := FALSE;
   // Movement.Request.MCMovement07WP := FALSE;
   // Movement.Request.MCMovement08WP := FALSE;
   // Movement.Request.MCMovement09WP := FALSE;
   // Movement.Request.MCMovement10WP := FALSE;
   // Movement.Request.MCMovement11WP := FALSE;
   // Movement.Request.MCMovement12WP := FALSE;
   // Movement.Request.MCMovement13WP := FALSE;
   // Movement.Request.MCMovement14WP := FALSE;
   // Movement.Request.MCMovement15WP := FALSE;
   // Movement.Request.MCMovement16WP := FALSE;
   // Movement.Request.MCMovement17WP := FALSE;
   // Movement.Request.MCMovement18WP := FALSE;
   // Movement.Request.MCMovement19WP := FALSE;
   // Movement.Request.MCMovement20WP := FALSE;
   // Movement.Request.MCMovement21WP := FALSE;
   // Movement.Request.MCMovement22WP := FALSE;
   // Movement.Request.MCMovement23WP := FALSE;
   // Movement.Request.MCMovement24WP := FALSE;
   // Movement.Request.MCMovement25WP := FALSE;
   // Movement.Request.MCMovement26WP := FALSE;
   // Movement.Request.MCMovement27WP := FALSE;
   // Movement.Request.MCMovement28WP := FALSE;
   // Movement.Request.MCMovement29WP := FALSE;
   // Movement.Request.MCMovement30WP := FALSE;
   // Movement.Request.MCMovement31WP := FALSE;
   // Movement.Request.MCMovement32WP := FALSE;
   // Movement.Request.MCMovement01BP := FALSE;
   // Movement.Request.MCMovement02BP := FALSE;
   // Movement.Request.MCMovement03BP := FALSE;
   // Movement.Request.MCMovement04BP := FALSE;
   // Movement.Request.MCMovement05BP := FALSE;
   // Movement.Request.MCMovement06BP := FALSE;
   // Movement.Request.MCMovement07BP := FALSE;
   // Movement.Request.MCMovement08BP := FALSE;
   // // 600 more start values not shown
END_TYPE

TYPE "UDT_Vacuum"
VERSION : 0.0
   STRUCT
      FLT_motor_protection : Bool;   // Störung: Der Versorgungsspanuung oder des Motorschutzes Motor
      FLT_min_level_oil : Bool;   // Störung: Der minimale Füllstand des Öls wurde unterschritten
      FLT_presure_reached : Bool;   // Störung: Der Vakuumdrucke wurde nicht erreicht
      FLT_filter : Bool;   // Störung: Der Luftfilter ist verschmutzt
      FLT_lock_start : Bool;   // Störung: Beim Einschalten des Vakuums ist die Wiederanlaufsperre noch aktiv
      Spare_0_5 : Bool;
      Spare_0_6 : Bool;
      Spare_0_7 : Bool;
      Flag_T_ON : Bool;   // Flankenhilfsmerker zum Ein- Ausschalten des Hydraulikmotors
      Request : Bool;   // Anforderung zum Einschalten des Vakuum- Motors
      Spare_1_2 : Bool;
      Spare_1_3 : Bool;
      Spare_1_4 : Bool;
      Motor_Stern : Bool;   // Ansteuerung des Hydraulikmotors 01 am Netz // in Stern
      Motor_Dreieck : Bool;   // Ansteuerung des Hydraulikmotors 01 im Dreieck
      Ready_and_okay : Bool;   // Die Vakuumpumpe läuft wunschgemäß
   END_STRUCT;
END_TYPE

